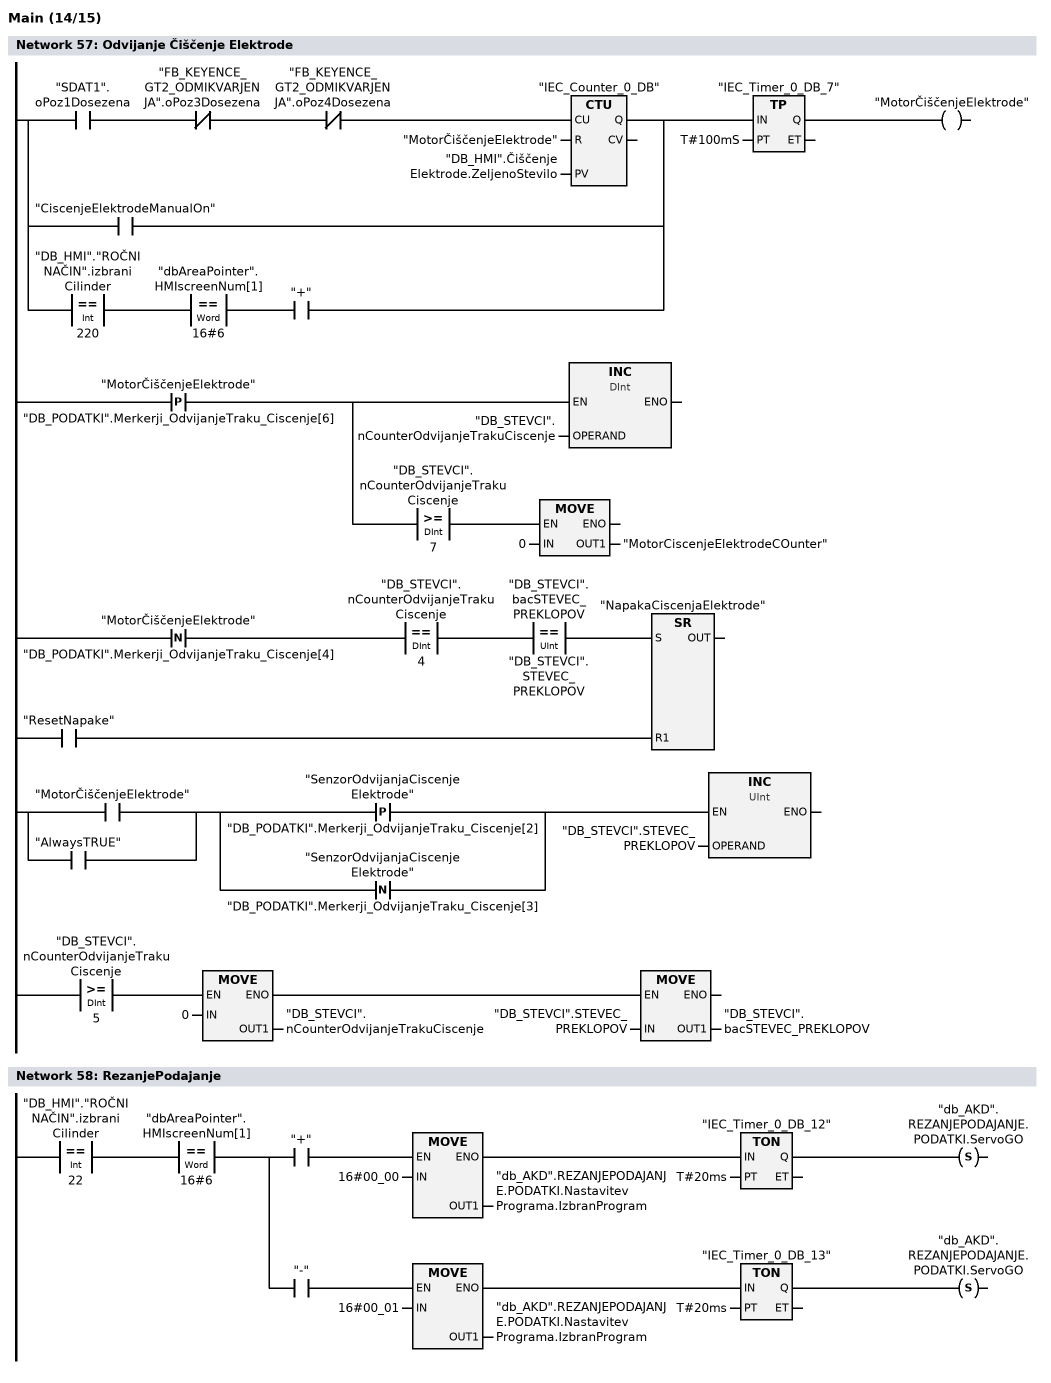
   "IEC_Counter_0_DB".CTU(CU := "SDAT1".oPoz1Dosezena AND NOT "FB_KEYENCE_GT2_ODMIKVARJENJA".oPoz3Dosezena AND NOT "FB_KEYENCE_GT2_ODMIKVARJENJA".oPoz4Dosezena,
                          R := "MotorČiščenjeElektrode",
                          PV := "DB_HMI".ČiščenjeElektrode.ZeljenoStevilo);
   "IEC_Timer_0_DB_7".TP(IN := "IEC_Counter_0_DB".Q OR "CiscenjeElektrodeManualOn" OR (("DB_HMI"."ROČNI NAČIN".izbraniCilinder = 220) AND ("dbAreaPointer".HMIscreenNum[1] = 16#6) AND "+"),
                         PT := T#100mS);
   "MotorČiščenjeElektrode" := "IEC_Timer_0_DB_7".Q;
   #_w1 := "MotorČiščenjeElektrode" AND NOT "DB_PODATKI".Merkerji_OdvijanjeTraku_Ciscenje[6];   // rising edge of "MotorČiščenjeElektrode"
   "DB_PODATKI".Merkerji_OdvijanjeTraku_Ciscenje[6] := "MotorČiščenjeElektrode";
   IF #_w1 THEN
       "DB_STEVCI".nCounterOdvijanjeTrakuCiscenje := "DB_STEVCI".nCounterOdvijanjeTrakuCiscenje + 1;
   END_IF;
   IF #_w1 AND ("DB_STEVCI".nCounterOdvijanjeTrakuCiscenje >= 7) THEN
       "MotorCiscenjeElektrodeCOunter" := 0;
   END_IF;
   #_w2 := NOT "MotorČiščenjeElektrode" AND "DB_PODATKI".Merkerji_OdvijanjeTraku_Ciscenje[4];   // falling edge of "MotorČiščenjeElektrode"
   "DB_PODATKI".Merkerji_OdvijanjeTraku_Ciscenje[4] := "MotorČiščenjeElektrode";
   IF #_w2 AND ("DB_STEVCI".nCounterOdvijanjeTrakuCiscenje = 4) AND ("DB_STEVCI".bacSTEVEC_PREKLOPOV = "DB_STEVCI".STEVEC_PREKLOPOV) THEN
       "NapakaCiscenjaElektrode" := TRUE;   // SR flip-flop
   END_IF;
   IF "ResetNapake" THEN "NapakaCiscenjaElektrode" := FALSE; END_IF;
   #_w3 := ("MotorČiščenjeElektrode" OR "AlwaysTRUE") AND "SenzorOdvijanjaCiscenjeElektrode" AND NOT "DB_PODATKI".Merkerji_OdvijanjeTraku_Ciscenje[2];   // rising edge of "SenzorOdvijanjaCiscenjeElektrode"
   "DB_PODATKI".Merkerji_OdvijanjeTraku_Ciscenje[2] := "SenzorOdvijanjaCiscenjeElektrode";
   #_w4 := ("MotorČiščenjeElektrode" OR "AlwaysTRUE") AND NOT "SenzorOdvijanjaCiscenjeElektrode" AND "DB_PODATKI".Merkerji_OdvijanjeTraku_Ciscenje[3];   // falling edge of "SenzorOdvijanjaCiscenjeElektrode"
   "DB_PODATKI".Merkerji_OdvijanjeTraku_Ciscenje[3] := "SenzorOdvijanjaCiscenjeElektrode";
   IF #_w3 OR #_w4 THEN "DB_STEVCI".STEVEC_PREKLOPOV := "DB_STEVCI".STEVEC_PREKLOPOV + 1; END_IF;
   #_w5 := "DB_STEVCI".nCounterOdvijanjeTrakuCiscenje >= 5;
   IF #_w5 THEN
       "DB_STEVCI".nCounterOdvijanjeTrakuCiscenje := 0;
       "DB_STEVCI".bacSTEVEC_PREKLOPOV := "DB_STEVCI".STEVEC_PREKLOPOV;
   END_IF;
END_REGION

REGION Network 58: RezanjePodajanje
   #_w1 := ("DB_HMI"."ROČNI NAČIN".izbraniCilinder = 22) AND ("dbAreaPointer".HMIscreenNum[1] = 16#6);
   #_w2 := #_w1 AND "+";
   IF #_w2 THEN "db_AKD".REZANJEPODAJANJE.PODATKI.NastavitevPrograma.IzbranProgram := 16#00_00; END_IF;
   "IEC_Timer_0_DB_12".TON(IN := #_w2, PT := T#20ms);
   IF "IEC_Timer_0_DB_12".Q THEN "db_AKD".REZANJEPODAJANJE.PODATKI.ServoGO := TRUE; END_IF;
   #_w3 := #_w1 AND "-";
   IF #_w3 THEN "db_AKD".REZANJEPODAJANJE.PODATKI.NastavitevPrograma.IzbranProgram := 16#00_01; END_IF;
   "IEC_Timer_0_DB_13".TON(IN := #_w3, PT := T#20ms);
   IF "IEC_Timer_0_DB_13".Q THEN "db_AKD".REZANJEPODAJANJE.PODATKI.ServoGO := TRUE; END_IF;
END_REGION

REGION Network 59: TEKOCI TRAK
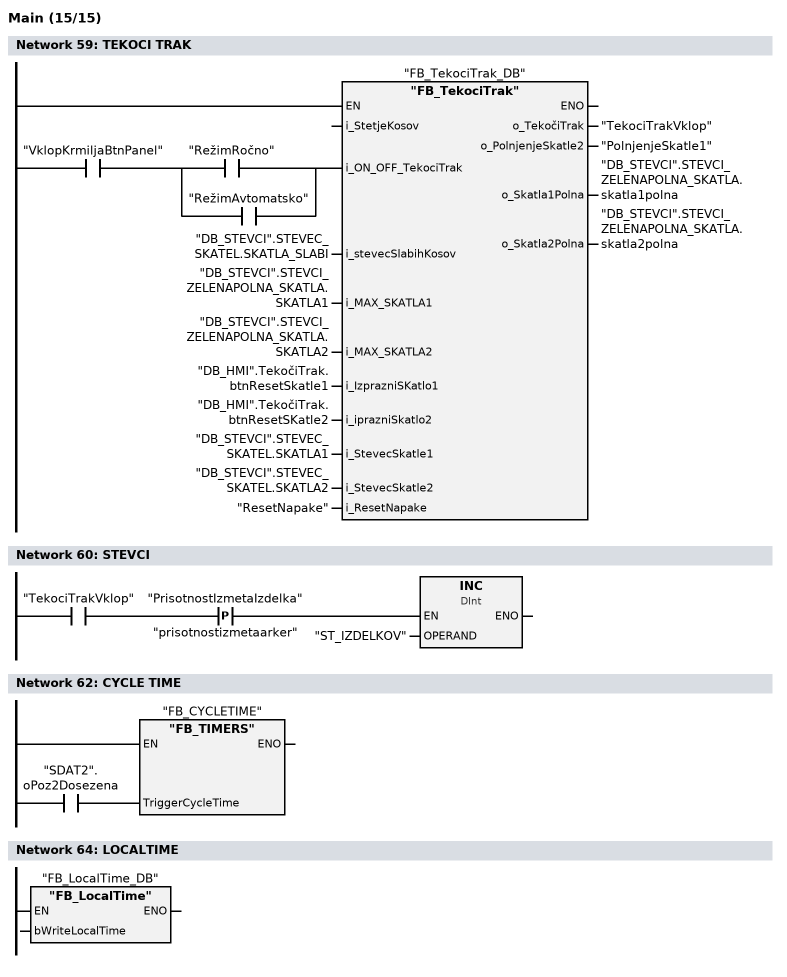
   RUNG wire#powerrail
      "FB_TekociTrak_DB"(i_ON_OFF_TekociTrak := wire#w2, i_StetjeKosov :=, i_stevecSlabihKosov := "DB_STEVCI".STEVEC_SKATEL.SKATLA_SLABI, i_MAX_SKATLA1 := "DB_STEVCI".STEVCI_ZELENAPOLNA_SKATLA.SKATLA1, i_MAX_SKATLA2 := "DB_STEVCI".STEVCI_ZELENAPOLNA_SKATLA.SKATLA2, i_IzprazniSKatlo1 := "DB_HMI".TekočiTrak.btnResetSkatle1, i_iprazniSkatlo2 := "DB_HMI".TekočiTrak.btnResetSKatle2, i_StevecSkatle1 := "DB_STEVCI".STEVEC_SKATEL.SKATLA1, i_StevecSkatle2 := "DB_STEVCI".STEVEC_SKATEL.SKATLA2, i_ResetNapake := "ResetNapake", o_TekočiTrak => "TekociTrakVklop", o_PolnjenjeSkatle2 => "PolnjenjeSkatle1", o_Skatla1Polna => "DB_STEVCI".STEVCI_ZELENAPOLNA_SKATLA.skatla1polna, o_Skatla2Polna => "DB_STEVCI".STEVCI_ZELENAPOLNA_SKATLA.skatla2polna)
   END_RUNG
   RUNG wire#powerrail
      Contact( "VklopKrmiljaBtnPanel" )
      wire#w1
      Contact( "RežimRočno" )
   END_RUNG wire#w2
   RUNG wire#w1
      Contact( "RežimAvtomatsko" )
   END_RUNG wire#w2
   // the same network as SCL:
   "FB_TekociTrak_DB"(i_ON_OFF_TekociTrak := "VklopKrmiljaBtnPanel" AND ("RežimRočno" OR "RežimAvtomatsko"),   // "FB_TekociTrak"
                      i_stevecSlabihKosov := "DB_STEVCI".STEVEC_SKATEL.SKATLA_SLABI,
                      i_MAX_SKATLA1 := "DB_STEVCI".STEVCI_ZELENAPOLNA_SKATLA.SKATLA1,
                      i_MAX_SKATLA2 := "DB_STEVCI".STEVCI_ZELENAPOLNA_SKATLA.SKATLA2,
                      i_IzprazniSKatlo1 := "DB_HMI".TekočiTrak.btnResetSkatle1,
                      i_iprazniSkatlo2 := "DB_HMI".TekočiTrak.btnResetSKatle2,
                      i_StevecSkatle1 := "DB_STEVCI".STEVEC_SKATEL.SKATLA1,
                      i_StevecSkatle2 := "DB_STEVCI".STEVEC_SKATEL.SKATLA2,
                      i_ResetNapake := "ResetNapake",
                      o_TekočiTrak => "TekociTrakVklop",
                      o_PolnjenjeSkatle2 => "PolnjenjeSkatle1",
                      o_Skatla1Polna => "DB_STEVCI".STEVCI_ZELENAPOLNA_SKATLA.skatla1polna,
                      o_Skatla2Polna => "DB_STEVCI".STEVCI_ZELENAPOLNA_SKATLA.skatla2polna);
END_REGION

REGION Network 60: STEVCI
   RUNG wire#powerrail
      Contact( "TekociTrakVklop" )
      P_Contact(operand := "PrisotnostIzmetaIzdelka", bit := "prisotnostizmetaarker")
      { S7_Templates := "DestType := DInt" } Inc( "ST_IZDELKOV" )
   END_RUNG
   // the same network as SCL:
   #_w1 := "TekociTrakVklop" AND "PrisotnostIzmetaIzdelka" AND NOT "prisotnostizmetaarker";   // rising edge of "PrisotnostIzmetaIzdelka"
   "prisotnostizmetaarker" := "PrisotnostIzmetaIzdelka";
   IF #_w1 THEN "ST_IZDELKOV" := "ST_IZDELKOV" + 1; END_IF;
END_REGION

REGION Network 62: CYCLE TIME
   RUNG wire#powerrail
      "FB_CYCLETIME"(TriggerCycleTime := wire#w1)
   END_RUNG
   RUNG wire#powerrail
      Contact( "SDAT2".oPoz2Dosezena )
   END_RUNG wire#w1
   // the same network as SCL:
   "FB_CYCLETIME"(TriggerCycleTime := "SDAT2".oPoz2Dosezena);   // "FB_TIMERS"
END_REGION

REGION Network 64: LOCALTIME
   RUNG wire#powerrail
      "FB_LocalTime_DB"(bWriteLocalTime :=)
   END_RUNG
   // the same network as SCL:
   "FB_LocalTime_DB"();   // "FB_LocalTime"
END_REGION
END_ORGANIZATION_BLOCK

ORGANIZATION_BLOCK "Startup"   // OB100, LAD, Startup
TITLE = "Complete Restart"
{ S7_Optimized_Access := 'TRUE' }
VERSION : 0.1
   VAR_INPUT
      LostRetentive : Bool;   // True if retentive data are lost
      LostRTC : Bool;   // True if date and time are lost
   END_VAR
BEGIN

REGION Network 1
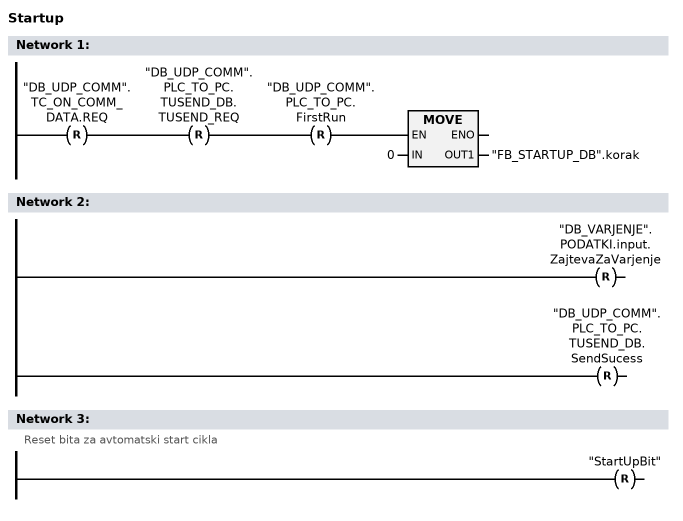
   RUNG wire#powerrail
      R_Coil( "DB_UDP_COMM".TC_ON_COMM_DATA.REQ )
      R_Coil( "DB_UDP_COMM".PLC_TO_PC.TUSEND_DB.TUSEND_REQ )
      R_Coil( "DB_UDP_COMM".PLC_TO_PC.FirstRun )
      Move(in := 0, out1 => "FB_STARTUP_DB".korak)
   END_RUNG
   // the same network as SCL:
   "DB_UDP_COMM".TC_ON_COMM_DATA.REQ := FALSE;
   "DB_UDP_COMM".PLC_TO_PC.TUSEND_DB.TUSEND_REQ := FALSE;
   "DB_UDP_COMM".PLC_TO_PC.FirstRun := FALSE;
   "FB_STARTUP_DB".korak := 0;
END_REGION

REGION Network 2
   RUNG wire#powerrail
      R_Coil( "DB_VARJENJE".PODATKI.input.ZajtevaZaVarjenje )
   END_RUNG
   RUNG wire#powerrail
      R_Coil( "DB_UDP_COMM".PLC_TO_PC.TUSEND_DB.SendSucess )
   END_RUNG
   // the same network as SCL:
   "DB_VARJENJE".PODATKI.input.ZajtevaZaVarjenje := FALSE;
   "DB_UDP_COMM".PLC_TO_PC.TUSEND_DB.SendSucess := FALSE;
END_REGION

REGION Network 3
   // Reset bita za avtomatski start cikla
   RUNG wire#powerrail
      R_Coil( "StartUpBit" )
   END_RUNG
   // the same network as SCL:
   "StartUpBit" := FALSE;
END_REGION
END_ORGANIZATION_BLOCK

ORGANIZATION_BLOCK "ProDiagOB"   // OB250, ProDiag_OB, ProgramCycle
TITLE = "Main Program Sweep (Cycle)"
{ S7_Optimized_Access := 'TRUE' }
VERSION : 0.1
   VAR_INPUT
      Initial_Call : Bool;   // Initial call of this OB
      Remanence : Bool;   // =True, if remanent data are available
   END_VAR
BEGIN

REGION Network 1
   CALL "Block_1", "Block_1_DB";
END_REGION
END_ORGANIZATION_BLOCK

// folder: FUNKCIJE/Funkcije

FUNCTION_BLOCK "FB_Lin_fun"   // FB9, LAD
TITLE = Izrčun izhoda po linearni funkciji
{ S7_Optimized_Access := 'TRUE' }
VERSION : 0.1
   VAR_INPUT
      I_PIW_real : Real := 0.0;
      I_x2 : Real := 100.0;
      I_x1 : Real := 0.0;
      I_y2 : Real := 100.0;
      I_y1 : Real := 0.0;
      I_napaka_signala : Real;
   END_VAR
   VAR_OUTPUT
      Q_izhod : Real := 0.0;
      Q_NAPAKA_signala : Bool;
   END_VAR
   VAR_TEMP
      Delta_y : Real;
      Delta_x : Real;
      K : Real;
      N : Real;
      Temp_real : Real;
   END_VAR
   VAR_TEMP   // added for the SCL form of the ladder/FBD networks
      _w1 : Bool;
   END_VAR
BEGIN

REGION Network 1: Izračun y2-y1 , x2-x1, k = (y2-y1) / (x2-x1)
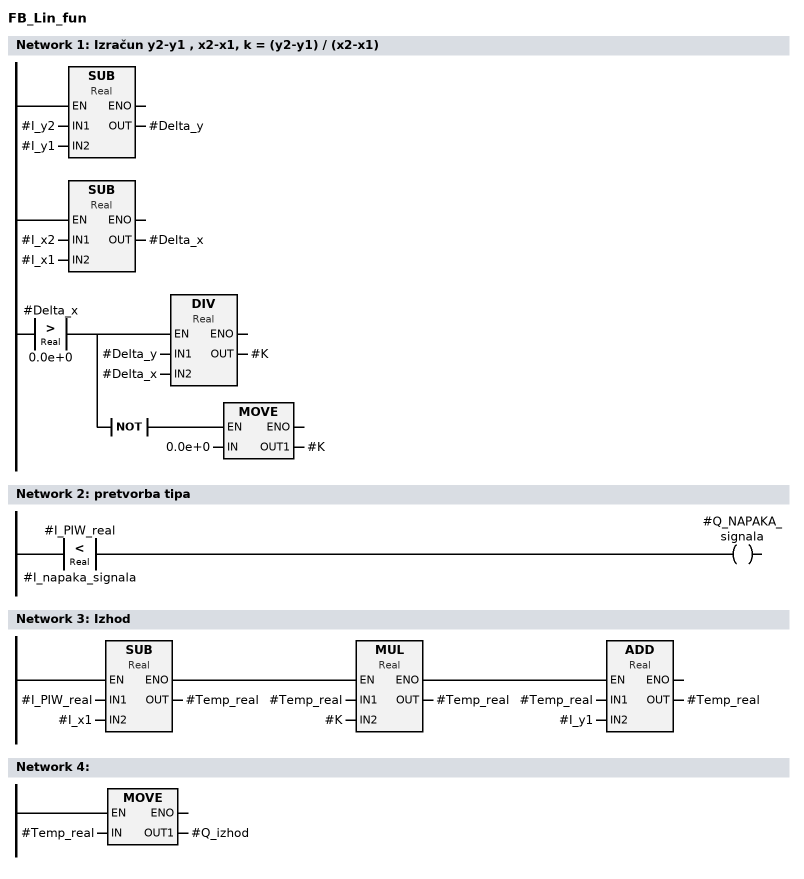
   RUNG wire#powerrail
      { S7_Templates := "SrcType := Real"; S7_GenerateENO := "TRUE" } Sub(in1 := #I_y2, in2 := #I_y1, out => #Delta_y)
   END_RUNG
   RUNG wire#powerrail
      { S7_Templates := "SrcType := Real"; S7_GenerateENO := "TRUE" } Sub(in1 := #I_x2, in2 := #I_x1, out => #Delta_x)
   END_RUNG
   RUNG wire#powerrail
      { S7_Templates := "SrcType := Real" } GT_Contact(in1 := #Delta_x, in2 := 0.0e+0)
      wire#w1
      { S7_Templates := "SrcType := Real"; S7_GenerateENO := "TRUE" } Div(in1 := #Delta_y, in2 := #Delta_x, out => #K)
   END_RUNG
   RUNG wire#w1
      Not()
      { S7_GenerateENO := "TRUE" } Move(in := 0.0e+0, out1 => #K)
   END_RUNG
   // the same network as SCL:
   #Delta_y := #I_y2 - #I_y1;
   #Delta_x := #I_x2 - #I_x1;
   #_w1 := #Delta_x > 0.0e+0;
   IF #_w1 THEN #K := #Delta_y / #Delta_x; END_IF;
   IF NOT #_w1 THEN #K := 0.0e+0; END_IF;
END_REGION

REGION Network 2: pretvorba tipa
   RUNG wire#powerrail
      { S7_Templates := "SrcType := Real" } LT_Contact(in1 := #I_PIW_real, in2 := #I_napaka_signala)
      Coil( #Q_NAPAKA_signala )
   END_RUNG
   // the same network as SCL:
   #Q_NAPAKA_signala := #I_PIW_real < #I_napaka_signala;
END_REGION

REGION Network 3: Izhod
   RUNG wire#powerrail
      { S7_Templates := "SrcType := Real"; S7_GenerateENO := "TRUE" } Sub(in1 := #I_PIW_real, in2 := #I_x1, out => #Temp_real)
      { S7_Templates := "SrcType := Real"; S7_GenerateENO := "TRUE" } Mul(in1 := #Temp_real, in2 := #K, out => #Temp_real)
      { S7_Templates := "SrcType := Real"; S7_GenerateENO := "TRUE" } Add(in1 := #Temp_real, in2 := #I_y1, out => #Temp_real)
   END_RUNG
   // the same network as SCL:
   // ENO of a box is taken as its EN; it also drops when the box reports an error
   #Temp_real := #I_PIW_real - #I_x1;
   #Temp_real := #Temp_real * #K;
   #Temp_real := #Temp_real + #I_y1;
END_REGION

REGION Network 4
   RUNG wire#powerrail
      { S7_GenerateENO := "TRUE" } Move(in := #Temp_real, out1 => #Q_izhod)
   END_RUNG
   // the same network as SCL:
   #Q_izhod := #Temp_real;
END_REGION
END_FUNCTION_BLOCK

FUNCTION_BLOCK "INT_TO_BOOL"   // FB10, SCL
{ S7_Optimized_Access := 'TRUE' }
VERSION : 0.1
   VAR_INPUT
      "INT" : Int;
   END_VAR
   VAR_OUTPUT
      BOOL_0 : Bool;
      BOOL_1 : Bool;
      BOOL_2 : Bool;
      BOOL_3 : Bool;
      BOOL_4 : Bool;
      BOOL_5 : Bool;
      BOOL_6 : Bool;
      BOOL_7 : Bool;
      BOOL_8 : Bool;
      BOOL_9 : Bool;
      BOOL_10 : Bool;
      BOOL_11 : Bool;
      BOOL_12 : Bool;
      BOOL_13 : Bool;
      BOOL_14 : Bool;
   END_VAR
   VAR
      INT_TEMP : Int;
   END_VAR
   VAR_TEMP
      statusna_beseda_temp : Int;
   END_VAR
BEGIN

   #INT_TEMP := SWAP(#INT);

   #statusna_beseda_temp := #INT_TEMP;
   #BOOL_0 := #statusna_beseda_temp.%X0;


   #statusna_beseda_temp := #INT_TEMP;
   #BOOL_1 := #statusna_beseda_temp.%X1;

   #statusna_beseda_temp := #INT_TEMP;
   #BOOL_2 := #statusna_beseda_temp.%X2;

   #statusna_beseda_temp := #INT_TEMP;
   #BOOL_3 := #statusna_beseda_temp.%X3;

   #statusna_beseda_temp := #INT_TEMP;
   #BOOL_4 := #statusna_beseda_temp.%X4;

   #statusna_beseda_temp := #INT_TEMP;
   #BOOL_5 := #statusna_beseda_temp.%X5;

   #statusna_beseda_temp := #INT_TEMP;
   #BOOL_6 := #statusna_beseda_temp.%X6;

   #statusna_beseda_temp := #INT_TEMP;
   #BOOL_7 := #statusna_beseda_temp.%X7;

   #statusna_beseda_temp := #INT_TEMP;
   #BOOL_8 := #statusna_beseda_temp.%X8;

   #statusna_beseda_temp := #INT_TEMP;
   #BOOL_9 := #statusna_beseda_temp.%X9;

   #statusna_beseda_temp := #INT_TEMP;
   #BOOL_10 := #statusna_beseda_temp.%X10;

   #statusna_beseda_temp := #INT_TEMP;
   #BOOL_11 := #statusna_beseda_temp.%X11;

   #statusna_beseda_temp := #INT_TEMP;
   #BOOL_12 := #statusna_beseda_temp.%X12;

   #statusna_beseda_temp := #INT_TEMP;
   #BOOL_13:= #statusna_beseda_temp.%X13;

   IF #statusna_beseda_temp > 0 THEN;
       #BOOL_14 := TRUE;

   ELSE
       #BOOL_14 := FALSE;
   END_IF;
END_FUNCTION_BLOCK

FUNCTION_BLOCK "Statistika_delovanja"   // FB32, LAD
{ S7_Optimized_Access := 'TRUE' }
VERSION : 0.1
   VAR_INPUT
      "Stevec serije" : DInt;
      "Stevec narejenih kosov" : DInt;
      Hitrost : DInt;
      faktor : DInt;
   END_VAR
   VAR
      Edge : Array[0..10] of Bool;
      "Minutni stevec" : Int;
      "Razlika kosov" : DInt;
      "Minute delovanja" : DInt;
      temp_ : DInt;
      "Preracun ure delovanja" : DInt;
      "Preracun minute delovanja" : DInt;
   END_VAR
   VAR_TEMP
      "temp 1" : DInt;
   END_VAR
   VAR_TEMP   // added for the SCL form of the ladder/FBD networks
      _w1 : Bool;
   END_VAR
BEGIN

REGION Network 2: izracun stevila kosov na minuto
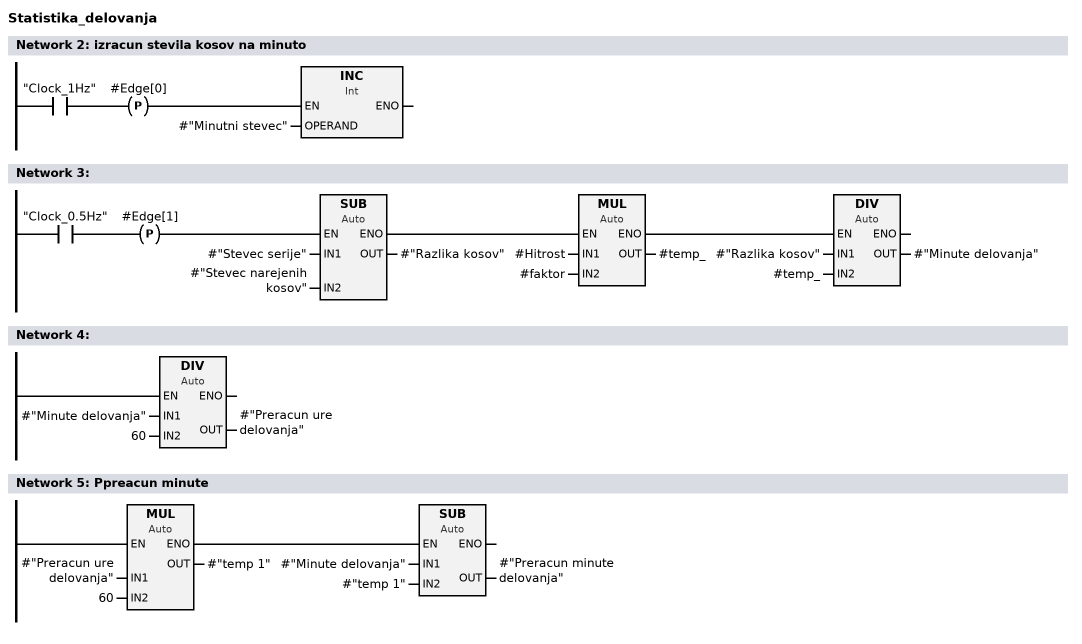
   RUNG wire#powerrail
      Contact( "Clock_1Hz" )
      P_Trig( #Edge[0] )
      { S7_Templates := "DestType := Int" } Inc( #"Minutni stevec" )
   END_RUNG
   // the same network as SCL:
   #_w1 := "Clock_1Hz" AND NOT #Edge[0];   // rising edge
   #Edge[0] := "Clock_1Hz";
   IF #_w1 THEN #"Minutni stevec" := #"Minutni stevec" + 1; END_IF;
END_REGION

REGION Network 3
   RUNG wire#powerrail
      Contact( "Clock_0.5Hz" )
      P_Trig( #Edge[1] )
      Sub(in1 := #"Stevec serije", in2 := #"Stevec narejenih kosov", out => #"Razlika kosov")
      Mul(in1 := #Hitrost, in2 := #faktor, out => #temp_)
      Div(in1 := #"Razlika kosov", in2 := #temp_, out => #"Minute delovanja")
   END_RUNG
   // the same network as SCL:
   #_w1 := "Clock_0.5Hz" AND NOT #Edge[1];   // rising edge
   #Edge[1] := "Clock_0.5Hz";
   IF #_w1 THEN
       #"Razlika kosov" := #"Stevec serije" - #"Stevec narejenih kosov";
       #temp_ := #Hitrost * #faktor;
       #"Minute delovanja" := #"Razlika kosov" / #temp_;
   END_IF;
END_REGION

REGION Network 4
   RUNG wire#powerrail
      Div(in1 := #"Minute delovanja", in2 := 60, out => #"Preracun ure delovanja")
   END_RUNG
   // the same network as SCL:
   #"Preracun ure delovanja" := #"Minute delovanja" / 60;
END_REGION

REGION Network 5: Ppreacun minute
   RUNG wire#powerrail
      Mul(in1 := #"Preracun ure delovanja", in2 := 60, out => #"temp 1")
      Sub(in1 := #"Minute delovanja", in2 := #"temp 1", out => #"Preracun minute delovanja")
   END_RUNG
   // the same network as SCL:
   #"temp 1" := #"Preracun ure delovanja" * 60;
   #"Preracun minute delovanja" := #"Minute delovanja" - #"temp 1";
END_REGION
END_FUNCTION_BLOCK

FUNCTION_BLOCK "FB_Alarms"   // FB124, LAD
TITLE = Alarm blok
{ S7_Optimized_Access := 'TRUE' }
AUTHOR : Andrej
VERSION : 0.1
// Alarm blok, za prozenje posameznih alarmov preko HMI
   VAR_INPUT
      I_FAULT_RESET : Bool;
      I_Alarm_0 : Bool;
      I_Alarm_1 : Bool;
      I_Alarm_2 : Bool;
      I_Alarm_3 : Bool;
      I_Alarm_4 : Bool;
      I_Alarm_5 : Bool;
      I_Alarm_6 : Bool;
      I_Alarm_7 : Bool;
      I_Alarm_8 : Bool;
      I_Alarm_9 : Bool;
      I_Alarm_10 : Bool;
      I_Alarm_11 : Bool;
      I_Alarm_12 : Bool;
      I_Alarm_13 : Bool;
      I_Alarm_14 : Bool;
      I_Alarm_15 : Bool;
      "Avtomatska potrditev alarma" : Bool;
   END_VAR
   VAR_OUTPUT
      Q_Alarm_word : Word;
      Q_General_fault : Bool;
   END_VAR
   VAR
      Temp_word : Word;
      I_Alarm_0_temp : Bool;
      I_Alarm_1_temp : Bool;
      I_Alarm_2_temp : Bool;
      I_Alarm_3_temp : Bool;
      I_Alarm_4_temp : Bool;
      I_Alarm_5_temp : Bool;
      I_Alarm_6_temp : Bool;
      I_Alarm_7_temp : Bool;
      I_Alarm_8_temp : Bool;
      I_Alarm_9_temp : Bool;
      I_Alarm_10_temp : Bool;
      I_Alarm_11_temp : Bool;
      I_Alarm_12_temp : Bool;
      I_Alarm_13_temp : Bool;
      I_Alarm_14_temp : Bool;
      I_Alarm_15_temp : Bool;
   END_VAR
BEGIN

REGION Network 1
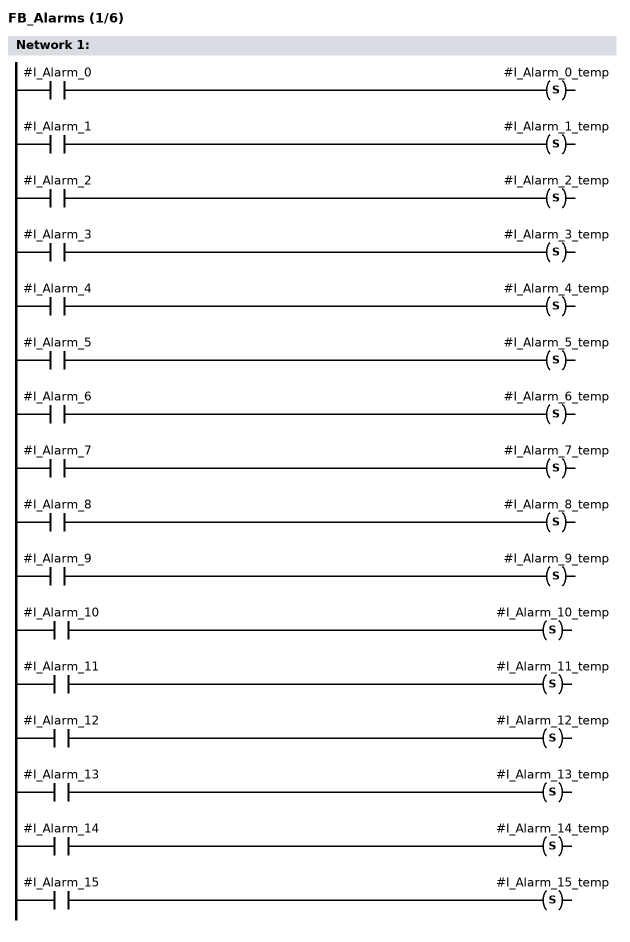
   RUNG wire#powerrail
      Contact( #I_Alarm_0 )
      S_Coil( #I_Alarm_0_temp )
   END_RUNG
   RUNG wire#powerrail
      Contact( #I_Alarm_1 )
      S_Coil( #I_Alarm_1_temp )
   END_RUNG
   RUNG wire#powerrail
      Contact( #I_Alarm_2 )
      S_Coil( #I_Alarm_2_temp )
   END_RUNG
   RUNG wire#powerrail
      Contact( #I_Alarm_3 )
      S_Coil( #I_Alarm_3_temp )
   END_RUNG
   RUNG wire#powerrail
      Contact( #I_Alarm_4 )
      S_Coil( #I_Alarm_4_temp )
   END_RUNG
   RUNG wire#powerrail
      Contact( #I_Alarm_5 )
      S_Coil( #I_Alarm_5_temp )
   END_RUNG
   RUNG wire#powerrail
      Contact( #I_Alarm_6 )
      S_Coil( #I_Alarm_6_temp )
   END_RUNG
   RUNG wire#powerrail
      Contact( #I_Alarm_7 )
      S_Coil( #I_Alarm_7_temp )
   END_RUNG
   RUNG wire#powerrail
      Contact( #I_Alarm_8 )
      S_Coil( #I_Alarm_8_temp )
   END_RUNG
   RUNG wire#powerrail
      Contact( #I_Alarm_9 )
      S_Coil( #I_Alarm_9_temp )
   END_RUNG
   RUNG wire#powerrail
      Contact( #I_Alarm_10 )
      S_Coil( #I_Alarm_10_temp )
   END_RUNG
   RUNG wire#powerrail
      Contact( #I_Alarm_11 )
      S_Coil( #I_Alarm_11_temp )
   END_RUNG
   RUNG wire#powerrail
      Contact( #I_Alarm_12 )
      S_Coil( #I_Alarm_12_temp )
   END_RUNG
   RUNG wire#powerrail
      Contact( #I_Alarm_13 )
      S_Coil( #I_Alarm_13_temp )
   END_RUNG
   RUNG wire#powerrail
      Contact( #I_Alarm_14 )
      S_Coil( #I_Alarm_14_temp )
   END_RUNG
   RUNG wire#powerrail
      Contact( #I_Alarm_15 )
      S_Coil( #I_Alarm_15_temp )
   END_RUNG
   // the same network as SCL:
   IF #I_Alarm_0 THEN #I_Alarm_0_temp := TRUE; END_IF;
   IF #I_Alarm_1 THEN #I_Alarm_1_temp := TRUE; END_IF;
   IF #I_Alarm_2 THEN #I_Alarm_2_temp := TRUE; END_IF;
   IF #I_Alarm_3 THEN #I_Alarm_3_temp := TRUE; END_IF;
   IF #I_Alarm_4 THEN #I_Alarm_4_temp := TRUE; END_IF;
   IF #I_Alarm_5 THEN #I_Alarm_5_temp := TRUE; END_IF;
   IF #I_Alarm_6 THEN #I_Alarm_6_temp := TRUE; END_IF;
   IF #I_Alarm_7 THEN #I_Alarm_7_temp := TRUE; END_IF;
   IF #I_Alarm_8 THEN #I_Alarm_8_temp := TRUE; END_IF;
   IF #I_Alarm_9 THEN #I_Alarm_9_temp := TRUE; END_IF;
   IF #I_Alarm_10 THEN #I_Alarm_10_temp := TRUE; END_IF;
   IF #I_Alarm_11 THEN #I_Alarm_11_temp := TRUE; END_IF;
   IF #I_Alarm_12 THEN #I_Alarm_12_temp := TRUE; END_IF;
   IF #I_Alarm_13 THEN #I_Alarm_13_temp := TRUE; END_IF;
   IF #I_Alarm_14 THEN #I_Alarm_14_temp := TRUE; END_IF;
   IF #I_Alarm_15 THEN #I_Alarm_15_temp := TRUE; END_IF;
END_REGION

REGION Network 2
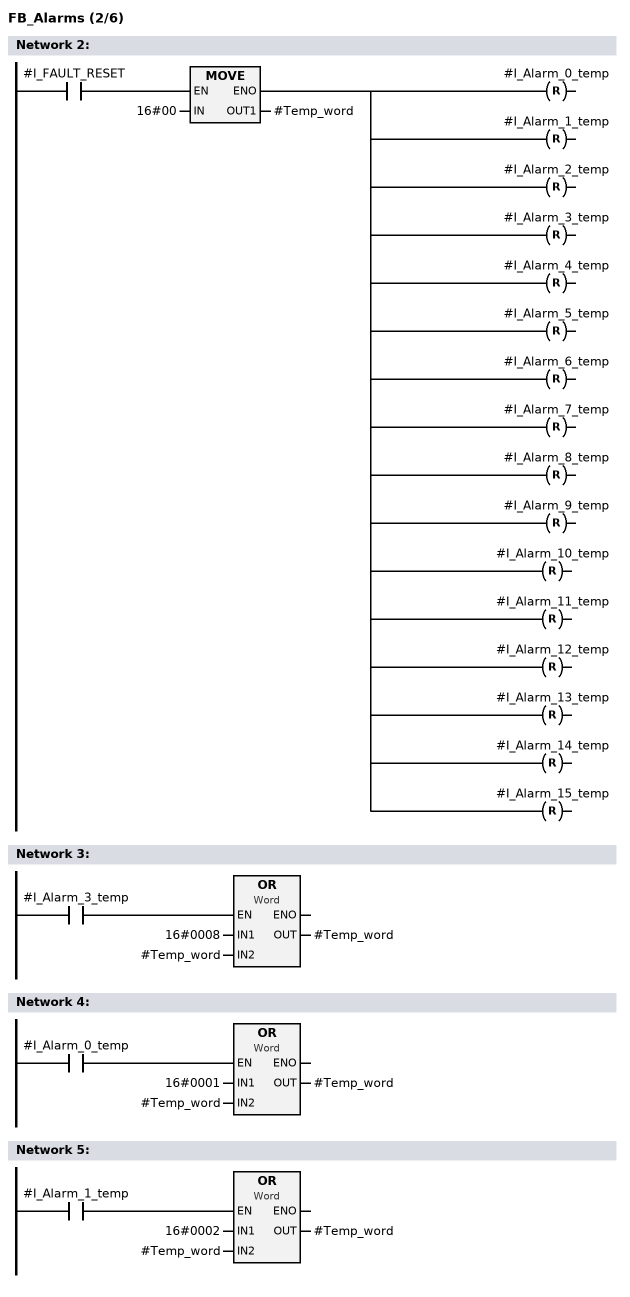
   RUNG wire#powerrail
      Contact( #I_FAULT_RESET )
      { S7_GenerateENO := "TRUE" } Move(in := 16#00, out1 => #Temp_word)
      wire#w1
      R_Coil( #I_Alarm_0_temp )
   END_RUNG
   RUNG wire#w1
      R_Coil( #I_Alarm_1_temp )
   END_RUNG
   RUNG wire#w1
      R_Coil( #I_Alarm_2_temp )
   END_RUNG
   RUNG wire#w1
      R_Coil( #I_Alarm_3_temp )
   END_RUNG
   RUNG wire#w1
      R_Coil( #I_Alarm_4_temp )
   END_RUNG
   RUNG wire#w1
      R_Coil( #I_Alarm_5_temp )
   END_RUNG
   RUNG wire#w1
      R_Coil( #I_Alarm_6_temp )
   END_RUNG
   RUNG wire#w1
      R_Coil( #I_Alarm_7_temp )
   END_RUNG
   RUNG wire#w1
      R_Coil( #I_Alarm_8_temp )
   END_RUNG
   RUNG wire#w1
      R_Coil( #I_Alarm_9_temp )
   END_RUNG
   RUNG wire#w1
      R_Coil( #I_Alarm_10_temp )
   END_RUNG
   RUNG wire#w1
      R_Coil( #I_Alarm_11_temp )
   END_RUNG
   RUNG wire#w1
      R_Coil( #I_Alarm_12_temp )
   END_RUNG
   RUNG wire#w1
      R_Coil( #I_Alarm_13_temp )
   END_RUNG
   RUNG wire#w1
      R_Coil( #I_Alarm_14_temp )
   END_RUNG
   RUNG wire#w1
      R_Coil( #I_Alarm_15_temp )
   END_RUNG
   // the same network as SCL:
   // ENO of a box is taken as its EN; it also drops when the box reports an error
   IF #I_FAULT_RESET THEN
       #Temp_word := 16#00;
       #I_Alarm_0_temp := FALSE;
       #I_Alarm_1_temp := FALSE;
       #I_Alarm_2_temp := FALSE;
       #I_Alarm_3_temp := FALSE;
       #I_Alarm_4_temp := FALSE;
       #I_Alarm_5_temp := FALSE;
       #I_Alarm_6_temp := FALSE;
       #I_Alarm_7_temp := FALSE;
       #I_Alarm_8_temp := FALSE;
       #I_Alarm_9_temp := FALSE;
       #I_Alarm_10_temp := FALSE;
       #I_Alarm_11_temp := FALSE;
       #I_Alarm_12_temp := FALSE;
       #I_Alarm_13_temp := FALSE;
       #I_Alarm_14_temp := FALSE;
       #I_Alarm_15_temp := FALSE;
   END_IF;
END_REGION

REGION Network 3
   IF #I_Alarm_3_temp THEN #Temp_word := 16#0008 OR #Temp_word; END_IF;
END_REGION

REGION Network 4
   IF #I_Alarm_0_temp THEN #Temp_word := 16#0001 OR #Temp_word; END_IF;
END_REGION

REGION Network 5
   IF #I_Alarm_1_temp THEN #Temp_word := 16#0002 OR #Temp_word; END_IF;
END_REGION

REGION Network 6
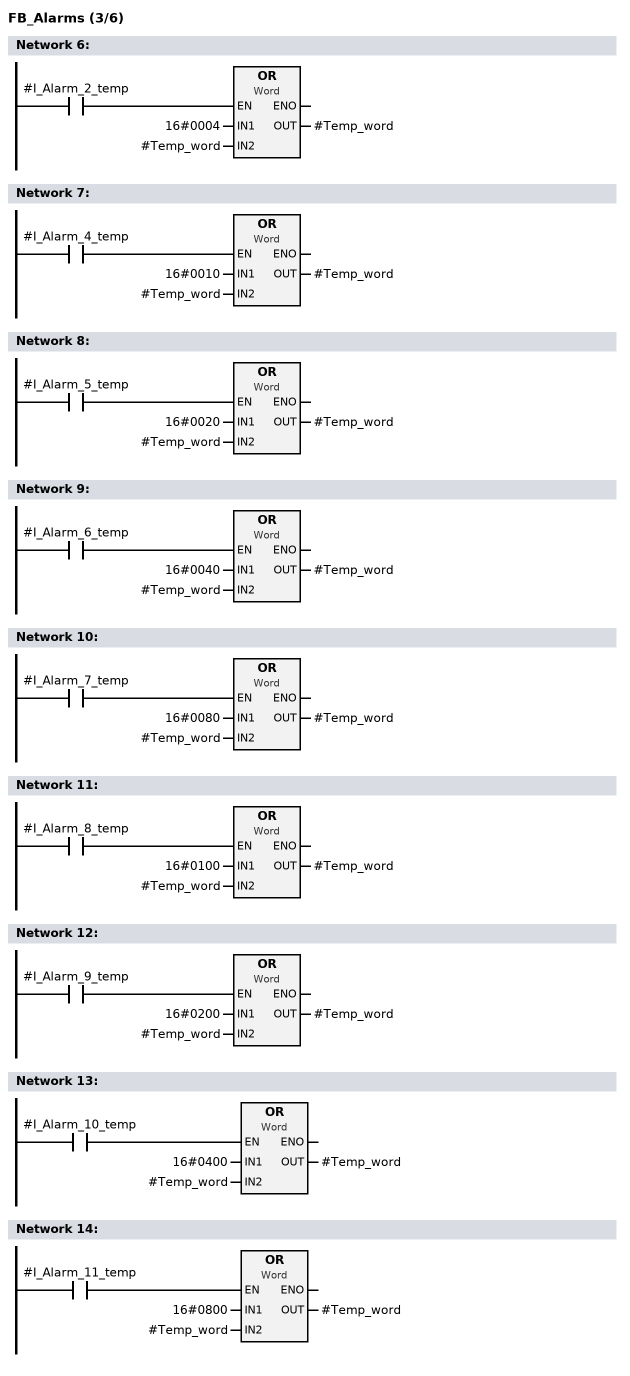
   IF #I_Alarm_2_temp THEN #Temp_word := 16#0004 OR #Temp_word; END_IF;
END_REGION

REGION Network 7
   IF #I_Alarm_4_temp THEN #Temp_word := 16#0010 OR #Temp_word; END_IF;
END_REGION

REGION Network 8
   IF #I_Alarm_5_temp THEN #Temp_word := 16#0020 OR #Temp_word; END_IF;
END_REGION

REGION Network 9
   IF #I_Alarm_6_temp THEN #Temp_word := 16#0040 OR #Temp_word; END_IF;
END_REGION

REGION Network 10
   IF #I_Alarm_7_temp THEN #Temp_word := 16#0080 OR #Temp_word; END_IF;
END_REGION

REGION Network 11
   IF #I_Alarm_8_temp THEN #Temp_word := 16#0100 OR #Temp_word; END_IF;
END_REGION

REGION Network 12
   IF #I_Alarm_9_temp THEN #Temp_word := 16#0200 OR #Temp_word; END_IF;
END_REGION

REGION Network 13
   IF #I_Alarm_10_temp THEN #Temp_word := 16#0400 OR #Temp_word; END_IF;
END_REGION

REGION Network 14
   IF #I_Alarm_11_temp THEN #Temp_word := 16#0800 OR #Temp_word; END_IF;
END_REGION

REGION Network 15
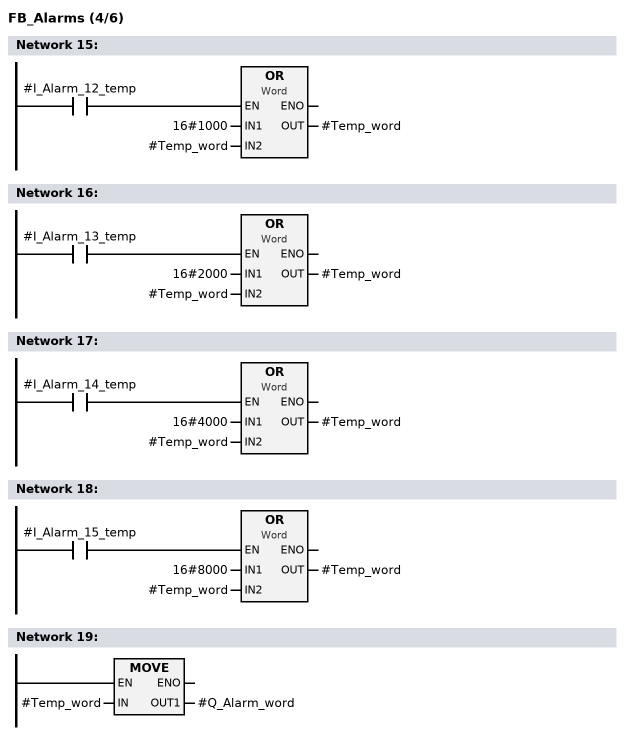
   IF #I_Alarm_12_temp THEN #Temp_word := 16#1000 OR #Temp_word; END_IF;
END_REGION

REGION Network 16
   IF #I_Alarm_13_temp THEN #Temp_word := 16#2000 OR #Temp_word; END_IF;
END_REGION

REGION Network 17
   IF #I_Alarm_14_temp THEN #Temp_word := 16#4000 OR #Temp_word; END_IF;
END_REGION

REGION Network 18
   IF #I_Alarm_15_temp THEN #Temp_word := 16#8000 OR #Temp_word; END_IF;
END_REGION

REGION Network 19
   RUNG wire#powerrail
      { S7_GenerateENO := "TRUE" } Move(in := #Temp_word, out1 => #Q_Alarm_word)
   END_RUNG
   // the same network as SCL:
   #Q_Alarm_word := #Temp_word;
END_REGION

REGION Network 20: General fault
